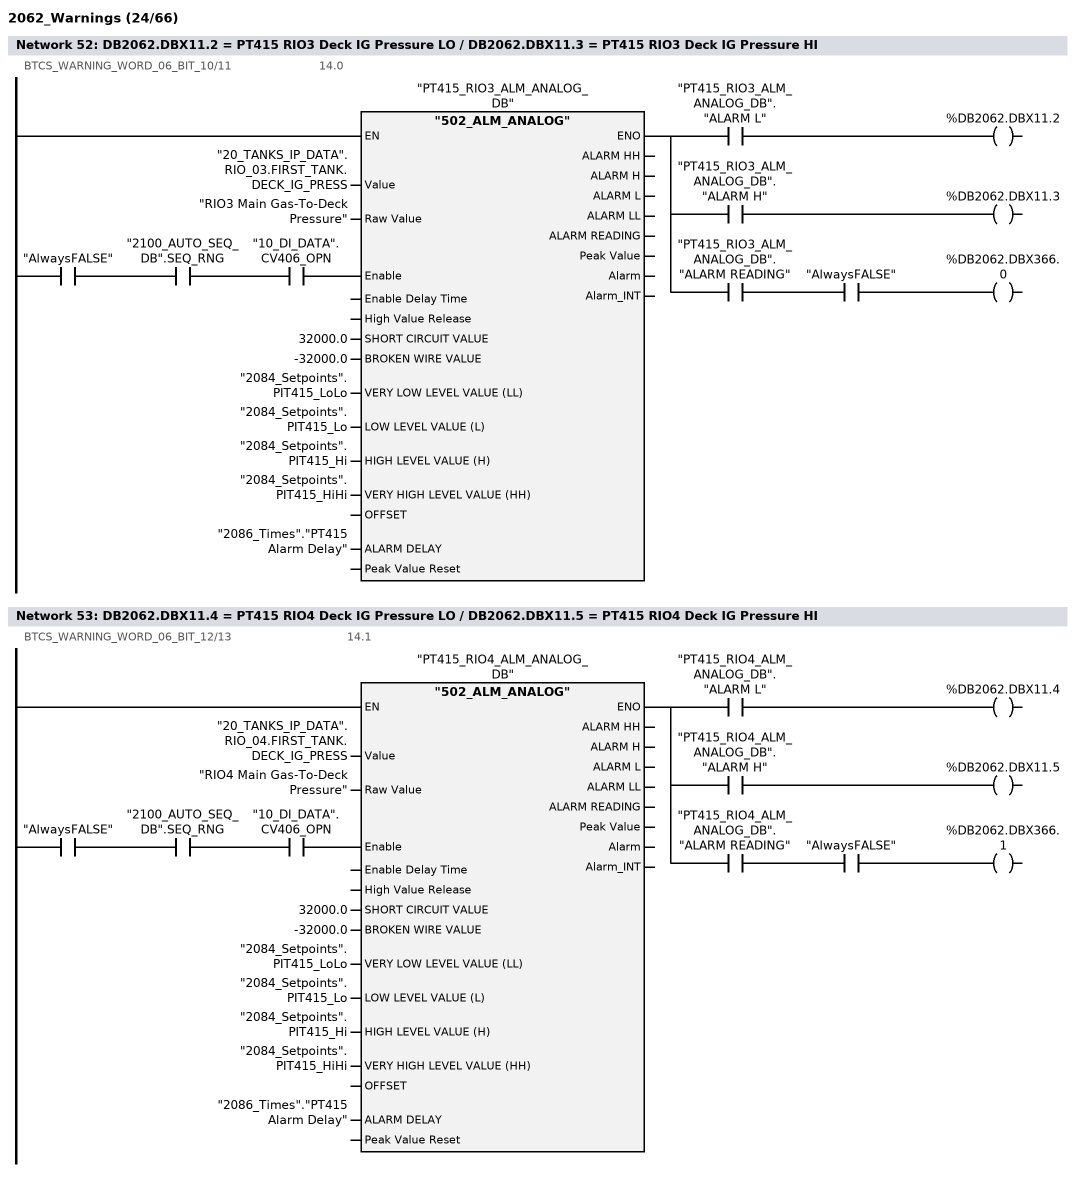
   RUNG wire#powerrail
      "PT415_RIO3_ALM_ANALOG_DB"(Enable := wire#w1, Value := "20_TANKS_IP_DATA".RIO_03.FIRST_TANK.DECK_IG_PRESS, "Raw Value" := "RIO3 Main Gas-To-Deck Pressure", "Enable Delay Time" :=, "High Value Release" :=, "SHORT CIRCUIT VALUE" := 32000.0, "BROKEN WIRE VALUE" := -32000.0, "VERY LOW LEVEL VALUE (LL)" := "2084_Setpoints".PIT415_LoLo, "LOW LEVEL VALUE (L)" := "2084_Setpoints".PIT415_Lo, "HIGH LEVEL VALUE (H)" := "2084_Setpoints".PIT415_Hi, "VERY HIGH LEVEL VALUE (HH)" := "2084_Setpoints".PIT415_HiHi, OFFSET :=, "ALARM DELAY" := "2086_Times"."PT415 Alarm Delay", "Peak Value Reset" :=, "ALARM HH" =>, "ALARM H" =>, "ALARM L" =>, "ALARM LL" =>, "ALARM READING" =>, "Peak Value" =>, Alarm =>, Alarm_INT =>)
      wire#w2
      Contact( "PT415_RIO3_ALM_ANALOG_DB"."ALARM L" )
      Coil( %DB2062.DBX11.2 )
   END_RUNG
   RUNG wire#powerrail
      Contact( "AlwaysFALSE" )
      Contact( "2100_AUTO_SEQ_DB".SEQ_RNG )
      Contact( "10_DI_DATA".CV406_OPN )
   END_RUNG wire#w1
   RUNG wire#w2
      Contact( "PT415_RIO3_ALM_ANALOG_DB"."ALARM H" )
      Coil( %DB2062.DBX11.3 )
   END_RUNG
   RUNG wire#w2
      Contact( "PT415_RIO3_ALM_ANALOG_DB"."ALARM READING" )
      Contact( "AlwaysFALSE" )
      Coil( %DB2062.DBX366.0 )
   END_RUNG
   // the same network as SCL:
   "PT415_RIO3_ALM_ANALOG_DB"(Value := "20_TANKS_IP_DATA".RIO_03.FIRST_TANK.DECK_IG_PRESS,   // "502_ALM_ANALOG"
                           "Raw Value" := "RIO3 Main Gas-To-Deck Pressure",
                           Enable := "AlwaysFALSE" AND "2100_AUTO_SEQ_DB".SEQ_RNG AND "10_DI_DATA".CV406_OPN,
                           "SHORT CIRCUIT VALUE" := 32000.0,
                           "BROKEN WIRE VALUE" := -32000.0,
                           "VERY LOW LEVEL VALUE (LL)" := "2084_Setpoints".PIT415_LoLo,
                           "LOW LEVEL VALUE (L)" := "2084_Setpoints".PIT415_Lo,
                           "HIGH LEVEL VALUE (H)" := "2084_Setpoints".PIT415_Hi,
                           "VERY HIGH LEVEL VALUE (HH)" := "2084_Setpoints".PIT415_HiHi,
                           "ALARM DELAY" := "2086_Times"."PT415 Alarm Delay",
                           ENO => #_w1);
   %DB2062.DBX11.2 := #_w1 AND "PT415_RIO3_ALM_ANALOG_DB"."ALARM L";
   %DB2062.DBX11.3 := #_w1 AND "PT415_RIO3_ALM_ANALOG_DB"."ALARM H";
   %DB2062.DBX366.0 := #_w1 AND "PT415_RIO3_ALM_ANALOG_DB"."ALARM READING" AND "AlwaysFALSE";
END_REGION

REGION Network 53: DB2062.DBX11.4 = PT415 RIO4 Deck IG Pressure LO / DB2062.DBX11.5 = PT415 RIO4 Deck IG Pressure HI
   // BTCS_WARNING_WORD_06_BIT_12/13                                 14.1
   RUNG wire#powerrail
      "PT415_RIO4_ALM_ANALOG_DB"(Enable := wire#w1, Value := "20_TANKS_IP_DATA".RIO_04.FIRST_TANK.DECK_IG_PRESS, "Raw Value" := "RIO4 Main Gas-To-Deck Pressure", "Enable Delay Time" :=, "High Value Release" :=, "SHORT CIRCUIT VALUE" := 32000.0, "BROKEN WIRE VALUE" := -32000.0, "VERY LOW LEVEL VALUE (LL)" := "2084_Setpoints".PIT415_LoLo, "LOW LEVEL VALUE (L)" := "2084_Setpoints".PIT415_Lo, "HIGH LEVEL VALUE (H)" := "2084_Setpoints".PIT415_Hi, "VERY HIGH LEVEL VALUE (HH)" := "2084_Setpoints".PIT415_HiHi, OFFSET :=, "ALARM DELAY" := "2086_Times"."PT415 Alarm Delay", "Peak Value Reset" :=, "ALARM HH" =>, "ALARM H" =>, "ALARM L" =>, "ALARM LL" =>, "ALARM READING" =>, "Peak Value" =>, Alarm =>, Alarm_INT =>)
      wire#w2
      Contact( "PT415_RIO4_ALM_ANALOG_DB"."ALARM L" )
      Coil( %DB2062.DBX11.4 )
   END_RUNG
   RUNG wire#powerrail
      Contact( "AlwaysFALSE" )
      Contact( "2100_AUTO_SEQ_DB".SEQ_RNG )
      Contact( "10_DI_DATA".CV406_OPN )
   END_RUNG wire#w1
   RUNG wire#w2
      Contact( "PT415_RIO4_ALM_ANALOG_DB"."ALARM H" )
      Coil( %DB2062.DBX11.5 )
   END_RUNG
   RUNG wire#w2
      Contact( "PT415_RIO4_ALM_ANALOG_DB"."ALARM READING" )
      Contact( "AlwaysFALSE" )
      Coil( %DB2062.DBX366.1 )
   END_RUNG
   // the same network as SCL:
   "PT415_RIO4_ALM_ANALOG_DB"(Value := "20_TANKS_IP_DATA".RIO_04.FIRST_TANK.DECK_IG_PRESS,   // "502_ALM_ANALOG"
                           "Raw Value" := "RIO4 Main Gas-To-Deck Pressure",
                           Enable := "AlwaysFALSE" AND "2100_AUTO_SEQ_DB".SEQ_RNG AND "10_DI_DATA".CV406_OPN,
                           "SHORT CIRCUIT VALUE" := 32000.0,
                           "BROKEN WIRE VALUE" := -32000.0,
                           "VERY LOW LEVEL VALUE (LL)" := "2084_Setpoints".PIT415_LoLo,
                           "LOW LEVEL VALUE (L)" := "2084_Setpoints".PIT415_Lo,
                           "HIGH LEVEL VALUE (H)" := "2084_Setpoints".PIT415_Hi,
                           "VERY HIGH LEVEL VALUE (HH)" := "2084_Setpoints".PIT415_HiHi,
                           "ALARM DELAY" := "2086_Times"."PT415 Alarm Delay",
                           ENO => #_w1);
   %DB2062.DBX11.4 := #_w1 AND "PT415_RIO4_ALM_ANALOG_DB"."ALARM L";
   %DB2062.DBX11.5 := #_w1 AND "PT415_RIO4_ALM_ANALOG_DB"."ALARM H";
   %DB2062.DBX366.1 := #_w1 AND "PT415_RIO4_ALM_ANALOG_DB"."ALARM READING" AND "AlwaysFALSE";
END_REGION

REGION Network 54: DB2062.DBX11.6 = PT415 RIO5 Deck IG Pressure LO / DB2062.DBX11.7 = PT415 RIO5 Deck IG Pressure HI
   // BTCS_WARNING_WORD_06_BIT_14/15                               14.2
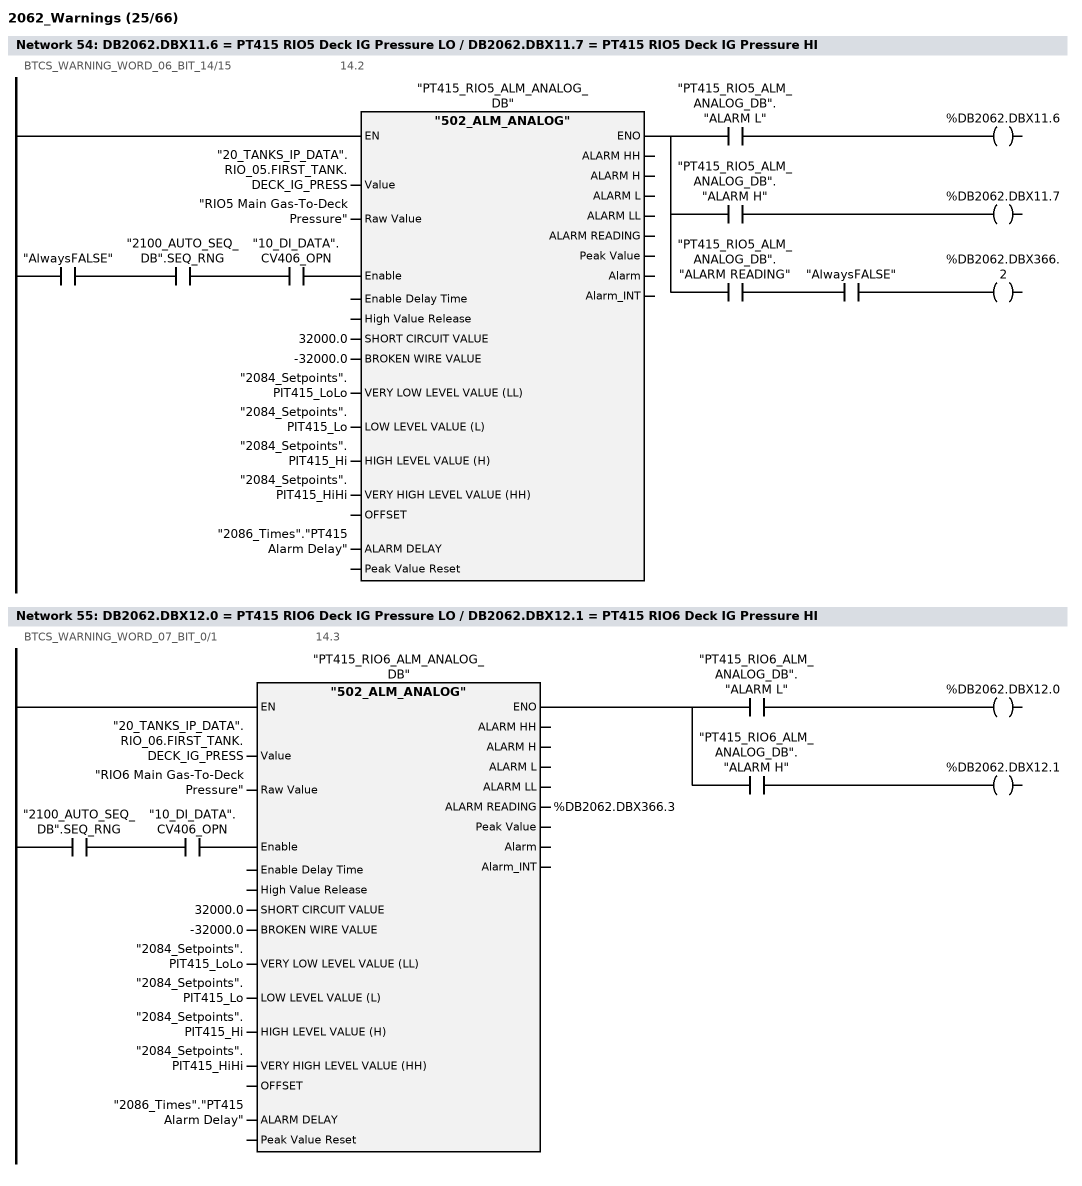
   RUNG wire#powerrail
      "PT415_RIO5_ALM_ANALOG_DB"(Enable := wire#w1, Value := "20_TANKS_IP_DATA".RIO_05.FIRST_TANK.DECK_IG_PRESS, "Raw Value" := "RIO5 Main Gas-To-Deck Pressure", "Enable Delay Time" :=, "High Value Release" :=, "SHORT CIRCUIT VALUE" := 32000.0, "BROKEN WIRE VALUE" := -32000.0, "VERY LOW LEVEL VALUE (LL)" := "2084_Setpoints".PIT415_LoLo, "LOW LEVEL VALUE (L)" := "2084_Setpoints".PIT415_Lo, "HIGH LEVEL VALUE (H)" := "2084_Setpoints".PIT415_Hi, "VERY HIGH LEVEL VALUE (HH)" := "2084_Setpoints".PIT415_HiHi, OFFSET :=, "ALARM DELAY" := "2086_Times"."PT415 Alarm Delay", "Peak Value Reset" :=, "ALARM HH" =>, "ALARM H" =>, "ALARM L" =>, "ALARM LL" =>, "ALARM READING" =>, "Peak Value" =>, Alarm =>, Alarm_INT =>)
      wire#w2
      Contact( "PT415_RIO5_ALM_ANALOG_DB"."ALARM L" )
      Coil( %DB2062.DBX11.6 )
   END_RUNG
   RUNG wire#powerrail
      Contact( "AlwaysFALSE" )
      Contact( "2100_AUTO_SEQ_DB".SEQ_RNG )
      Contact( "10_DI_DATA".CV406_OPN )
   END_RUNG wire#w1
   RUNG wire#w2
      Contact( "PT415_RIO5_ALM_ANALOG_DB"."ALARM H" )
      Coil( %DB2062.DBX11.7 )
   END_RUNG
   RUNG wire#w2
      Contact( "PT415_RIO5_ALM_ANALOG_DB"."ALARM READING" )
      Contact( "AlwaysFALSE" )
      Coil( %DB2062.DBX366.2 )
   END_RUNG
   // the same network as SCL:
   "PT415_RIO5_ALM_ANALOG_DB"(Value := "20_TANKS_IP_DATA".RIO_05.FIRST_TANK.DECK_IG_PRESS,   // "502_ALM_ANALOG"
                           "Raw Value" := "RIO5 Main Gas-To-Deck Pressure",
                           Enable := "AlwaysFALSE" AND "2100_AUTO_SEQ_DB".SEQ_RNG AND "10_DI_DATA".CV406_OPN,
                           "SHORT CIRCUIT VALUE" := 32000.0,
                           "BROKEN WIRE VALUE" := -32000.0,
                           "VERY LOW LEVEL VALUE (LL)" := "2084_Setpoints".PIT415_LoLo,
                           "LOW LEVEL VALUE (L)" := "2084_Setpoints".PIT415_Lo,
                           "HIGH LEVEL VALUE (H)" := "2084_Setpoints".PIT415_Hi,
                           "VERY HIGH LEVEL VALUE (HH)" := "2084_Setpoints".PIT415_HiHi,
                           "ALARM DELAY" := "2086_Times"."PT415 Alarm Delay",
                           ENO => #_w1);
   %DB2062.DBX11.6 := #_w1 AND "PT415_RIO5_ALM_ANALOG_DB"."ALARM L";
   %DB2062.DBX11.7 := #_w1 AND "PT415_RIO5_ALM_ANALOG_DB"."ALARM H";
   %DB2062.DBX366.2 := #_w1 AND "PT415_RIO5_ALM_ANALOG_DB"."ALARM READING" AND "AlwaysFALSE";
END_REGION

REGION Network 55: DB2062.DBX12.0 = PT415 RIO6 Deck IG Pressure LO / DB2062.DBX12.1 = PT415 RIO6 Deck IG Pressure HI
   // BTCS_WARNING_WORD_07_BIT_0/1                            14.3
   RUNG wire#powerrail
      "PT415_RIO6_ALM_ANALOG_DB"(Enable := wire#w1, Value := "20_TANKS_IP_DATA".RIO_06.FIRST_TANK.DECK_IG_PRESS, "Raw Value" := "RIO6 Main Gas-To-Deck Pressure", "Enable Delay Time" :=, "High Value Release" :=, "SHORT CIRCUIT VALUE" := 32000.0, "BROKEN WIRE VALUE" := -32000.0, "VERY LOW LEVEL VALUE (LL)" := "2084_Setpoints".PIT415_LoLo, "LOW LEVEL VALUE (L)" := "2084_Setpoints".PIT415_Lo, "HIGH LEVEL VALUE (H)" := "2084_Setpoints".PIT415_Hi, "VERY HIGH LEVEL VALUE (HH)" := "2084_Setpoints".PIT415_HiHi, OFFSET :=, "ALARM DELAY" := "2086_Times"."PT415 Alarm Delay", "Peak Value Reset" :=, "ALARM HH" =>, "ALARM H" =>, "ALARM L" =>, "ALARM LL" =>, "ALARM READING" => %DB2062.DBX366.3, "Peak Value" =>, Alarm =>, Alarm_INT =>)
      wire#w2
      Contact( "PT415_RIO6_ALM_ANALOG_DB"."ALARM L" )
      Coil( %DB2062.DBX12.0 )
   END_RUNG
   RUNG wire#powerrail
      Contact( "2100_AUTO_SEQ_DB".SEQ_RNG )
      Contact( "10_DI_DATA".CV406_OPN )
   END_RUNG wire#w1
   RUNG wire#w2
      Contact( "PT415_RIO6_ALM_ANALOG_DB"."ALARM H" )
      Coil( %DB2062.DBX12.1 )
   END_RUNG
   // the same network as SCL:
   "PT415_RIO6_ALM_ANALOG_DB"(Value := "20_TANKS_IP_DATA".RIO_06.FIRST_TANK.DECK_IG_PRESS,   // "502_ALM_ANALOG"
                           "Raw Value" := "RIO6 Main Gas-To-Deck Pressure",
                           Enable := "2100_AUTO_SEQ_DB".SEQ_RNG AND "10_DI_DATA".CV406_OPN,
                           "SHORT CIRCUIT VALUE" := 32000.0,
                           "BROKEN WIRE VALUE" := -32000.0,
                           "VERY LOW LEVEL VALUE (LL)" := "2084_Setpoints".PIT415_LoLo,
                           "LOW LEVEL VALUE (L)" := "2084_Setpoints".PIT415_Lo,
                           "HIGH LEVEL VALUE (H)" := "2084_Setpoints".PIT415_Hi,
                           "VERY HIGH LEVEL VALUE (HH)" := "2084_Setpoints".PIT415_HiHi,
                           "ALARM DELAY" := "2086_Times"."PT415 Alarm Delay",
                           "ALARM READING" => %DB2062.DBX366.3,
                           ENO => #_w1);
   %DB2062.DBX12.0 := #_w1 AND "PT415_RIO6_ALM_ANALOG_DB"."ALARM L";
   %DB2062.DBX12.1 := #_w1 AND "PT415_RIO6_ALM_ANALOG_DB"."ALARM H";
END_REGION

REGION Network 56: DB2062.DBX14.0 = PT415 RIO7 Deck IG Pressure LO / DB2062.DBX14.1 = PT415 RIO7 Deck IG Pressure HI
   // BTCS_WARNING_WORD_08_BIT_0/1                        14.4
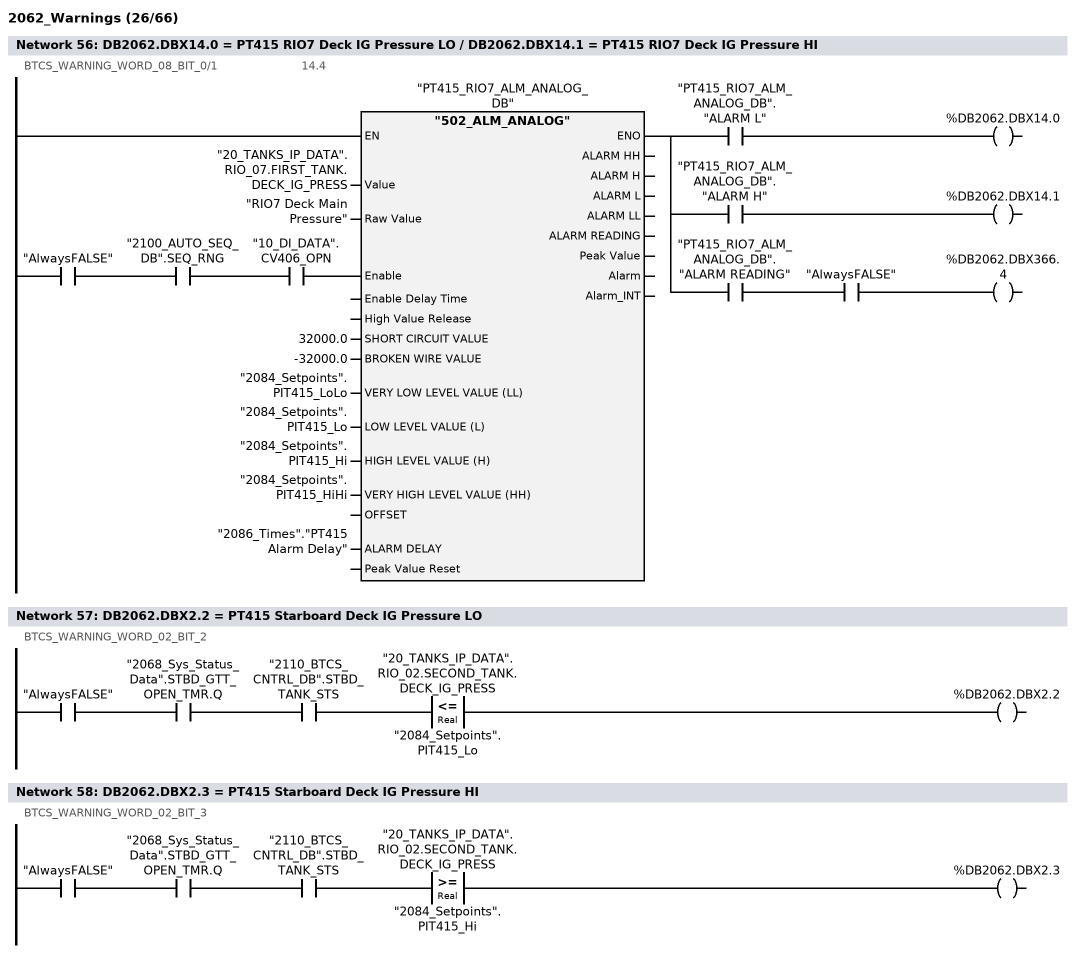
   RUNG wire#powerrail
      "PT415_RIO7_ALM_ANALOG_DB"(Enable := wire#w1, Value := "20_TANKS_IP_DATA".RIO_07.FIRST_TANK.DECK_IG_PRESS, "Raw Value" := "RIO7 Deck Main Pressure", "Enable Delay Time" :=, "High Value Release" :=, "SHORT CIRCUIT VALUE" := 32000.0, "BROKEN WIRE VALUE" := -32000.0, "VERY LOW LEVEL VALUE (LL)" := "2084_Setpoints".PIT415_LoLo, "LOW LEVEL VALUE (L)" := "2084_Setpoints".PIT415_Lo, "HIGH LEVEL VALUE (H)" := "2084_Setpoints".PIT415_Hi, "VERY HIGH LEVEL VALUE (HH)" := "2084_Setpoints".PIT415_HiHi, OFFSET :=, "ALARM DELAY" := "2086_Times"."PT415 Alarm Delay", "Peak Value Reset" :=, "ALARM HH" =>, "ALARM H" =>, "ALARM L" =>, "ALARM LL" =>, "ALARM READING" =>, "Peak Value" =>, Alarm =>, Alarm_INT =>)
      wire#w2
      Contact( "PT415_RIO7_ALM_ANALOG_DB"."ALARM L" )
      Coil( %DB2062.DBX14.0 )
   END_RUNG
   RUNG wire#powerrail
      Contact( "AlwaysFALSE" )
      Contact( "2100_AUTO_SEQ_DB".SEQ_RNG )
      Contact( "10_DI_DATA".CV406_OPN )
   END_RUNG wire#w1
   RUNG wire#w2
      Contact( "PT415_RIO7_ALM_ANALOG_DB"."ALARM H" )
      Coil( %DB2062.DBX14.1 )
   END_RUNG
   RUNG wire#w2
      Contact( "PT415_RIO7_ALM_ANALOG_DB"."ALARM READING" )
      Contact( "AlwaysFALSE" )
      Coil( %DB2062.DBX366.4 )
   END_RUNG
   // the same network as SCL:
   "PT415_RIO7_ALM_ANALOG_DB"(Value := "20_TANKS_IP_DATA".RIO_07.FIRST_TANK.DECK_IG_PRESS,   // "502_ALM_ANALOG"
                           "Raw Value" := "RIO7 Deck Main Pressure",
                           Enable := "AlwaysFALSE" AND "2100_AUTO_SEQ_DB".SEQ_RNG AND "10_DI_DATA".CV406_OPN,
                           "SHORT CIRCUIT VALUE" := 32000.0,
                           "BROKEN WIRE VALUE" := -32000.0,
                           "VERY LOW LEVEL VALUE (LL)" := "2084_Setpoints".PIT415_LoLo,
                           "LOW LEVEL VALUE (L)" := "2084_Setpoints".PIT415_Lo,
                           "HIGH LEVEL VALUE (H)" := "2084_Setpoints".PIT415_Hi,
                           "VERY HIGH LEVEL VALUE (HH)" := "2084_Setpoints".PIT415_HiHi,
                           "ALARM DELAY" := "2086_Times"."PT415 Alarm Delay",
                           ENO => #_w1);
   %DB2062.DBX14.0 := #_w1 AND "PT415_RIO7_ALM_ANALOG_DB"."ALARM L";
   %DB2062.DBX14.1 := #_w1 AND "PT415_RIO7_ALM_ANALOG_DB"."ALARM H";
   %DB2062.DBX366.4 := #_w1 AND "PT415_RIO7_ALM_ANALOG_DB"."ALARM READING" AND "AlwaysFALSE";
END_REGION

REGION Network 57: DB2062.DBX2.2 = PT415 Starboard Deck IG Pressure LO
   // BTCS_WARNING_WORD_02_BIT_2
   RUNG wire#powerrail
      Contact( "AlwaysFALSE" )
      Contact( "2068_Sys_Status_Data".STBD_GTT_OPEN_TMR.Q )
      Contact( "2110_BTCS_CNTRL_DB".STBD_TANK_STS )
      { S7_Templates := "SrcType := Real" } LE_Contact(in1 := "20_TANKS_IP_DATA".RIO_02.SECOND_TANK.DECK_IG_PRESS, in2 := "2084_Setpoints".PIT415_Lo)
      Coil( %DB2062.DBX2.2 )
   END_RUNG
   // the same network as SCL:
   %DB2062.DBX2.2 := "AlwaysFALSE" AND "2068_Sys_Status_Data".STBD_GTT_OPEN_TMR.Q AND "2110_BTCS_CNTRL_DB".STBD_TANK_STS AND ("20_TANKS_IP_DATA".RIO_02.SECOND_TANK.DECK_IG_PRESS <= "2084_Setpoints".PIT415_Lo);
END_REGION

REGION Network 58: DB2062.DBX2.3 = PT415 Starboard Deck IG Pressure HI
   // BTCS_WARNING_WORD_02_BIT_3
   RUNG wire#powerrail
      Contact( "AlwaysFALSE" )
      Contact( "2068_Sys_Status_Data".STBD_GTT_OPEN_TMR.Q )
      Contact( "2110_BTCS_CNTRL_DB".STBD_TANK_STS )
      { S7_Templates := "SrcType := Real" } GE_Contact(in1 := "20_TANKS_IP_DATA".RIO_02.SECOND_TANK.DECK_IG_PRESS, in2 := "2084_Setpoints".PIT415_Hi)
      Coil( %DB2062.DBX2.3 )
   END_RUNG
   // the same network as SCL:
   %DB2062.DBX2.3 := "AlwaysFALSE" AND "2068_Sys_Status_Data".STBD_GTT_OPEN_TMR.Q AND "2110_BTCS_CNTRL_DB".STBD_TANK_STS AND ("20_TANKS_IP_DATA".RIO_02.SECOND_TANK.DECK_IG_PRESS >= "2084_Setpoints".PIT415_Hi);
END_REGION

REGION Network 60: DB2062.DBX12.2/3 = PIT424 RIO1 Tank Pressure LO/HI
   // BTCS_WARNING_WORD_07_BIT_2/3                          14.5
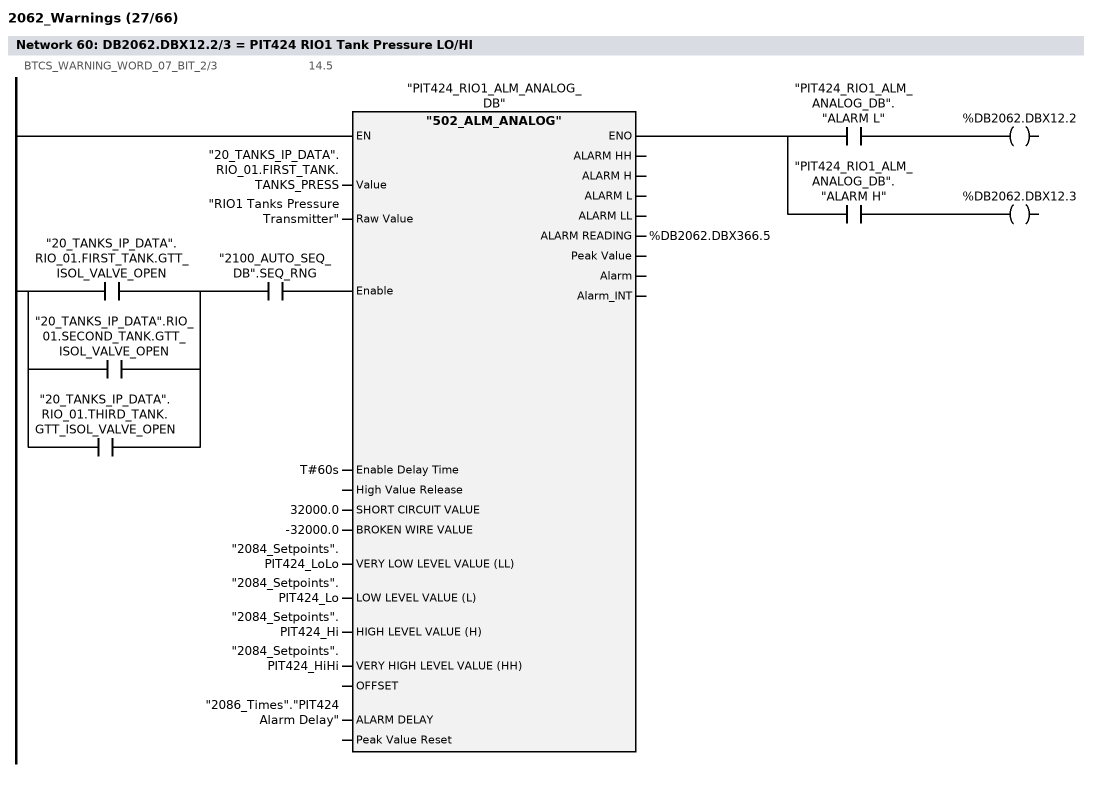
   RUNG wire#powerrail
      "PIT424_RIO1_ALM_ANALOG_DB"(Enable := wire#w2, Value := "20_TANKS_IP_DATA".RIO_01.FIRST_TANK.TANKS_PRESS, "Raw Value" := "RIO1 Tanks Pressure Transmitter", "Enable Delay Time" := T#60s, "High Value Release" :=, "SHORT CIRCUIT VALUE" := 32000.0, "BROKEN WIRE VALUE" := -32000.0, "VERY LOW LEVEL VALUE (LL)" := "2084_Setpoints".PIT424_LoLo, "LOW LEVEL VALUE (L)" := "2084_Setpoints".PIT424_Lo, "HIGH LEVEL VALUE (H)" := "2084_Setpoints".PIT424_Hi, "VERY HIGH LEVEL VALUE (HH)" := "2084_Setpoints".PIT424_HiHi, OFFSET :=, "ALARM DELAY" := "2086_Times"."PIT424 Alarm Delay", "Peak Value Reset" :=, "ALARM HH" =>, "ALARM H" =>, "ALARM L" =>, "ALARM LL" =>, "ALARM READING" => %DB2062.DBX366.5, "Peak Value" =>, Alarm =>, Alarm_INT =>)
      wire#w3
      Contact( "PIT424_RIO1_ALM_ANALOG_DB"."ALARM L" )
      Coil( %DB2062.DBX12.2 )
   END_RUNG
   RUNG wire#powerrail
      Contact( "20_TANKS_IP_DATA".RIO_01.FIRST_TANK.GTT_ISOL_VALVE_OPEN )
      wire#w1
      Contact( "2100_AUTO_SEQ_DB".SEQ_RNG )
   END_RUNG wire#w2
   RUNG wire#powerrail
      Contact( "20_TANKS_IP_DATA".RIO_01.SECOND_TANK.GTT_ISOL_VALVE_OPEN )
   END_RUNG wire#w1
   RUNG wire#powerrail
      Contact( "20_TANKS_IP_DATA".RIO_01.THIRD_TANK.GTT_ISOL_VALVE_OPEN )
   END_RUNG wire#w1
   RUNG wire#w3
      Contact( "PIT424_RIO1_ALM_ANALOG_DB"."ALARM H" )
      Coil( %DB2062.DBX12.3 )
   END_RUNG
   // the same network as SCL:
   "PIT424_RIO1_ALM_ANALOG_DB"(Value := "20_TANKS_IP_DATA".RIO_01.FIRST_TANK.TANKS_PRESS,   // "502_ALM_ANALOG"
                           "Raw Value" := "RIO1 Tanks Pressure Transmitter",
                           Enable := ("20_TANKS_IP_DATA".RIO_01.FIRST_TANK.GTT_ISOL_VALVE_OPEN OR "20_TANKS_IP_DATA".RIO_01.SECOND_TANK.GTT_ISOL_VALVE_OPEN OR "20_TANKS_IP_DATA".RIO_01.THIRD_TANK.GTT_ISOL_VALVE_OPEN) AND "2100_AUTO_SEQ_DB".SEQ_RNG,
                           "Enable Delay Time" := T#60s,
                           "SHORT CIRCUIT VALUE" := 32000.0,
                           "BROKEN WIRE VALUE" := -32000.0,
                           "VERY LOW LEVEL VALUE (LL)" := "2084_Setpoints".PIT424_LoLo,
                           "LOW LEVEL VALUE (L)" := "2084_Setpoints".PIT424_Lo,
                           "HIGH LEVEL VALUE (H)" := "2084_Setpoints".PIT424_Hi,
                           "VERY HIGH LEVEL VALUE (HH)" := "2084_Setpoints".PIT424_HiHi,
                           "ALARM DELAY" := "2086_Times"."PIT424 Alarm Delay",
                           "ALARM READING" => %DB2062.DBX366.5,
                           ENO => #_w1);
   %DB2062.DBX12.2 := #_w1 AND "PIT424_RIO1_ALM_ANALOG_DB"."ALARM L";
   %DB2062.DBX12.3 := #_w1 AND "PIT424_RIO1_ALM_ANALOG_DB"."ALARM H";
END_REGION

REGION Network 61: DB2062.DBX2.4/5 = PIT424 RIO2 Tank Pressure LO/HI
   // BTCS_WARNING_WORD_02_BIT_4                       14.6
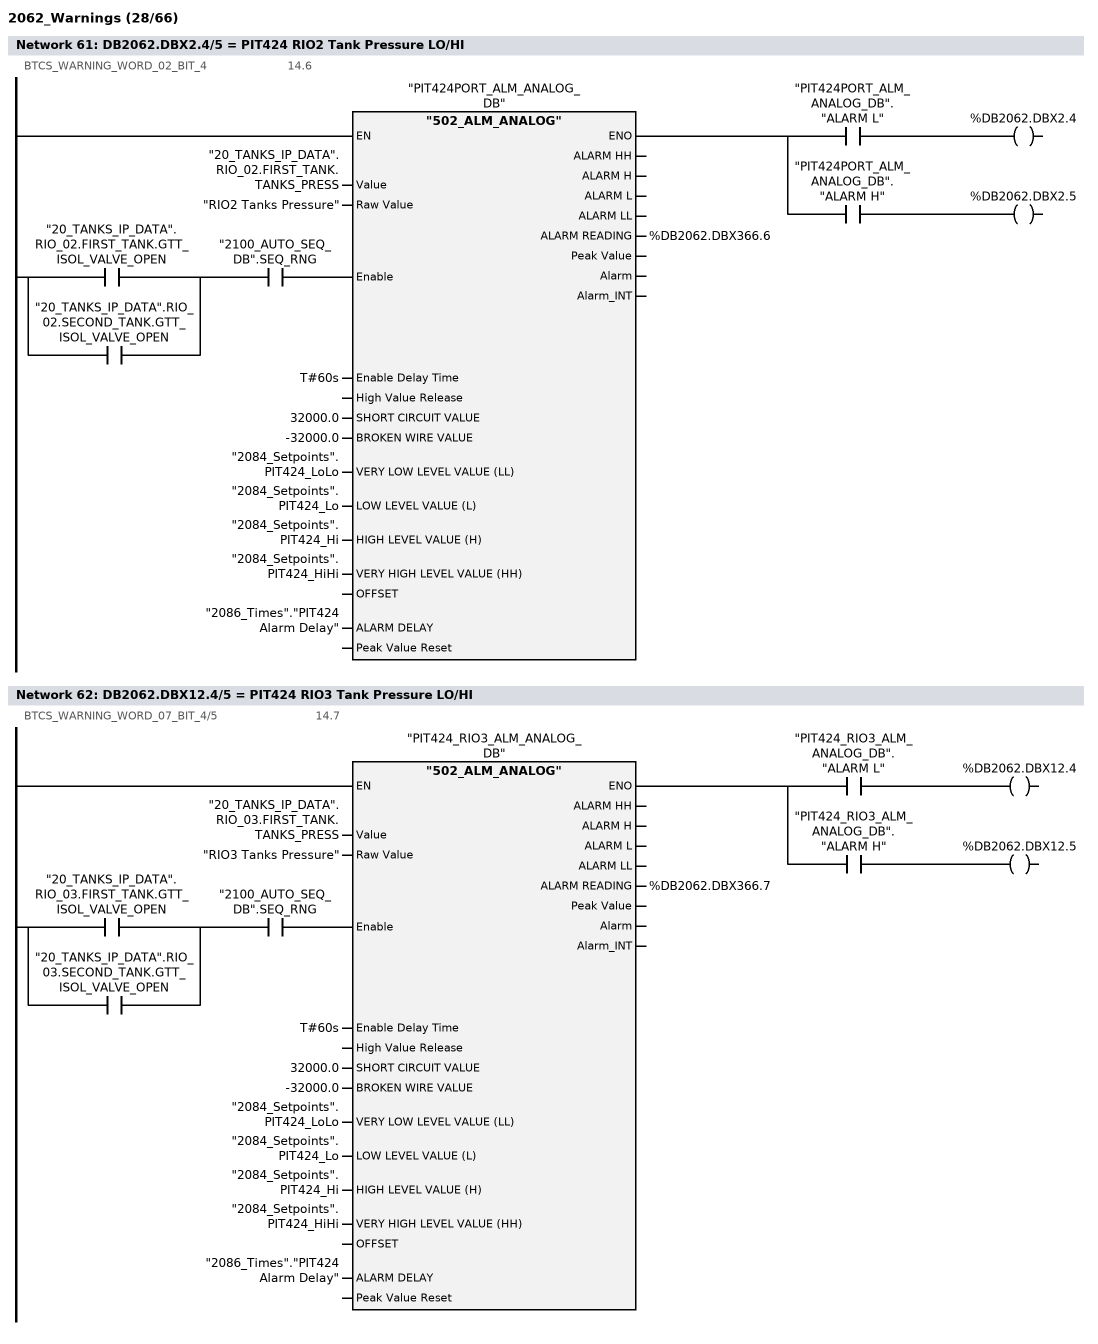
   RUNG wire#powerrail
      "PIT424PORT_ALM_ANALOG_DB"(Enable := wire#w2, Value := "20_TANKS_IP_DATA".RIO_02.FIRST_TANK.TANKS_PRESS, "Raw Value" := "RIO2 Tanks Pressure", "Enable Delay Time" := T#60s, "High Value Release" :=, "SHORT CIRCUIT VALUE" := 32000.0, "BROKEN WIRE VALUE" := -32000.0, "VERY LOW LEVEL VALUE (LL)" := "2084_Setpoints".PIT424_LoLo, "LOW LEVEL VALUE (L)" := "2084_Setpoints".PIT424_Lo, "HIGH LEVEL VALUE (H)" := "2084_Setpoints".PIT424_Hi, "VERY HIGH LEVEL VALUE (HH)" := "2084_Setpoints".PIT424_HiHi, OFFSET :=, "ALARM DELAY" := "2086_Times"."PIT424 Alarm Delay", "Peak Value Reset" :=, "ALARM HH" =>, "ALARM H" =>, "ALARM L" =>, "ALARM LL" =>, "ALARM READING" => %DB2062.DBX366.6, "Peak Value" =>, Alarm =>, Alarm_INT =>)
      wire#w3
      Contact( "PIT424PORT_ALM_ANALOG_DB"."ALARM L" )
      Coil( %DB2062.DBX2.4 )
   END_RUNG
   RUNG wire#powerrail
      Contact( "20_TANKS_IP_DATA".RIO_02.FIRST_TANK.GTT_ISOL_VALVE_OPEN )
      wire#w1
      Contact( "2100_AUTO_SEQ_DB".SEQ_RNG )
   END_RUNG wire#w2
   RUNG wire#powerrail
      Contact( "20_TANKS_IP_DATA".RIO_02.SECOND_TANK.GTT_ISOL_VALVE_OPEN )
   END_RUNG wire#w1
   RUNG wire#w3
      Contact( "PIT424PORT_ALM_ANALOG_DB"."ALARM H" )
      Coil( %DB2062.DBX2.5 )
   END_RUNG
   // the same network as SCL:
   "PIT424PORT_ALM_ANALOG_DB"(Value := "20_TANKS_IP_DATA".RIO_02.FIRST_TANK.TANKS_PRESS,   // "502_ALM_ANALOG"
                           "Raw Value" := "RIO2 Tanks Pressure",
                           Enable := ("20_TANKS_IP_DATA".RIO_02.FIRST_TANK.GTT_ISOL_VALVE_OPEN OR "20_TANKS_IP_DATA".RIO_02.SECOND_TANK.GTT_ISOL_VALVE_OPEN) AND "2100_AUTO_SEQ_DB".SEQ_RNG,
                           "Enable Delay Time" := T#60s,
                           "SHORT CIRCUIT VALUE" := 32000.0,
                           "BROKEN WIRE VALUE" := -32000.0,
                           "VERY LOW LEVEL VALUE (LL)" := "2084_Setpoints".PIT424_LoLo,
                           "LOW LEVEL VALUE (L)" := "2084_Setpoints".PIT424_Lo,
                           "HIGH LEVEL VALUE (H)" := "2084_Setpoints".PIT424_Hi,
                           "VERY HIGH LEVEL VALUE (HH)" := "2084_Setpoints".PIT424_HiHi,
                           "ALARM DELAY" := "2086_Times"."PIT424 Alarm Delay",
                           "ALARM READING" => %DB2062.DBX366.6,
                           ENO => #_w1);
   %DB2062.DBX2.4 := #_w1 AND "PIT424PORT_ALM_ANALOG_DB"."ALARM L";
   %DB2062.DBX2.5 := #_w1 AND "PIT424PORT_ALM_ANALOG_DB"."ALARM H";
END_REGION

REGION Network 62: DB2062.DBX12.4/5 = PIT424 RIO3 Tank Pressure LO/HI
   // BTCS_WARNING_WORD_07_BIT_4/5                            14.7
   RUNG wire#powerrail
      "PIT424_RIO3_ALM_ANALOG_DB"(Enable := wire#w2, Value := "20_TANKS_IP_DATA".RIO_03.FIRST_TANK.TANKS_PRESS, "Raw Value" := "RIO3 Tanks Pressure", "Enable Delay Time" := T#60s, "High Value Release" :=, "SHORT CIRCUIT VALUE" := 32000.0, "BROKEN WIRE VALUE" := -32000.0, "VERY LOW LEVEL VALUE (LL)" := "2084_Setpoints".PIT424_LoLo, "LOW LEVEL VALUE (L)" := "2084_Setpoints".PIT424_Lo, "HIGH LEVEL VALUE (H)" := "2084_Setpoints".PIT424_Hi, "VERY HIGH LEVEL VALUE (HH)" := "2084_Setpoints".PIT424_HiHi, OFFSET :=, "ALARM DELAY" := "2086_Times"."PIT424 Alarm Delay", "Peak Value Reset" :=, "ALARM HH" =>, "ALARM H" =>, "ALARM L" =>, "ALARM LL" =>, "ALARM READING" => %DB2062.DBX366.7, "Peak Value" =>, Alarm =>, Alarm_INT =>)
      wire#w3
      Contact( "PIT424_RIO3_ALM_ANALOG_DB"."ALARM L" )
      Coil( %DB2062.DBX12.4 )
   END_RUNG
   RUNG wire#powerrail
      Contact( "20_TANKS_IP_DATA".RIO_03.FIRST_TANK.GTT_ISOL_VALVE_OPEN )
      wire#w1
      Contact( "2100_AUTO_SEQ_DB".SEQ_RNG )
   END_RUNG wire#w2
   RUNG wire#powerrail
      Contact( "20_TANKS_IP_DATA".RIO_03.SECOND_TANK.GTT_ISOL_VALVE_OPEN )
   END_RUNG wire#w1
   RUNG wire#w3
      Contact( "PIT424_RIO3_ALM_ANALOG_DB"."ALARM H" )
      Coil( %DB2062.DBX12.5 )
   END_RUNG
   // the same network as SCL:
   "PIT424_RIO3_ALM_ANALOG_DB"(Value := "20_TANKS_IP_DATA".RIO_03.FIRST_TANK.TANKS_PRESS,   // "502_ALM_ANALOG"
                           "Raw Value" := "RIO3 Tanks Pressure",
                           Enable := ("20_TANKS_IP_DATA".RIO_03.FIRST_TANK.GTT_ISOL_VALVE_OPEN OR "20_TANKS_IP_DATA".RIO_03.SECOND_TANK.GTT_ISOL_VALVE_OPEN) AND "2100_AUTO_SEQ_DB".SEQ_RNG,
                           "Enable Delay Time" := T#60s,
                           "SHORT CIRCUIT VALUE" := 32000.0,
                           "BROKEN WIRE VALUE" := -32000.0,
                           "VERY LOW LEVEL VALUE (LL)" := "2084_Setpoints".PIT424_LoLo,
                           "LOW LEVEL VALUE (L)" := "2084_Setpoints".PIT424_Lo,
                           "HIGH LEVEL VALUE (H)" := "2084_Setpoints".PIT424_Hi,
                           "VERY HIGH LEVEL VALUE (HH)" := "2084_Setpoints".PIT424_HiHi,
                           "ALARM DELAY" := "2086_Times"."PIT424 Alarm Delay",
                           "ALARM READING" => %DB2062.DBX366.7,
                           ENO => #_w1);
   %DB2062.DBX12.4 := #_w1 AND "PIT424_RIO3_ALM_ANALOG_DB"."ALARM L";
   %DB2062.DBX12.5 := #_w1 AND "PIT424_RIO3_ALM_ANALOG_DB"."ALARM H";
END_REGION

REGION Network 63: DB2062.DBX12.6/7 = PIT424 RIO4 Tank Pressure LO/HI
   // BTCS_WARNING_WORD_07_BIT_6/7                           14.8
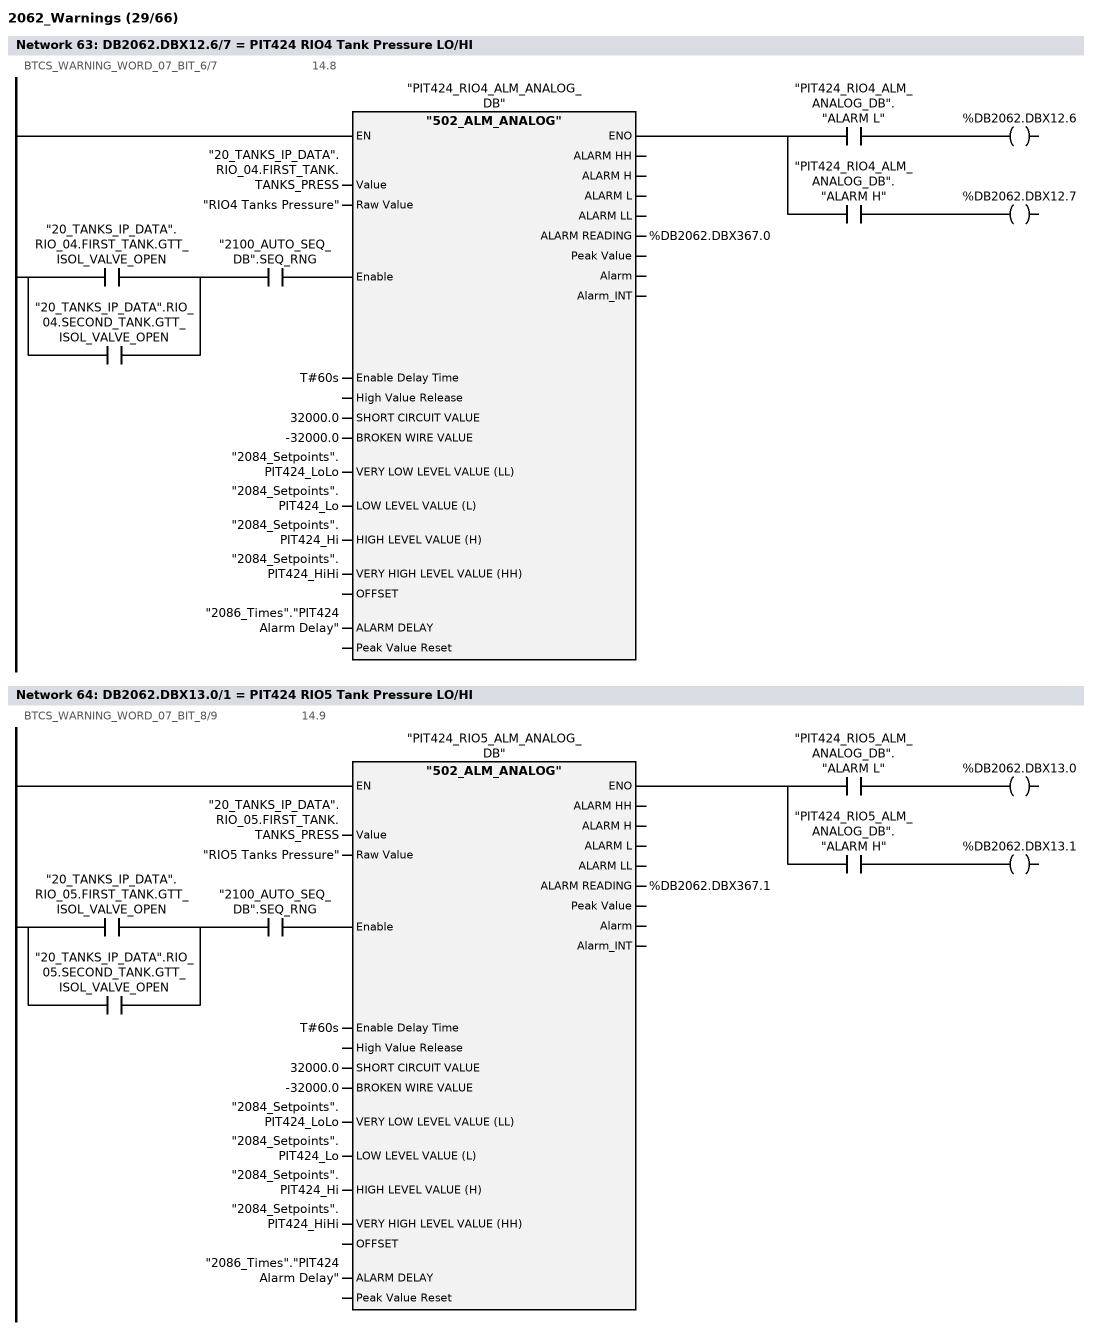
   RUNG wire#powerrail
      "PIT424_RIO4_ALM_ANALOG_DB"(Enable := wire#w2, Value := "20_TANKS_IP_DATA".RIO_04.FIRST_TANK.TANKS_PRESS, "Raw Value" := "RIO4 Tanks Pressure", "Enable Delay Time" := T#60s, "High Value Release" :=, "SHORT CIRCUIT VALUE" := 32000.0, "BROKEN WIRE VALUE" := -32000.0, "VERY LOW LEVEL VALUE (LL)" := "2084_Setpoints".PIT424_LoLo, "LOW LEVEL VALUE (L)" := "2084_Setpoints".PIT424_Lo, "HIGH LEVEL VALUE (H)" := "2084_Setpoints".PIT424_Hi, "VERY HIGH LEVEL VALUE (HH)" := "2084_Setpoints".PIT424_HiHi, OFFSET :=, "ALARM DELAY" := "2086_Times"."PIT424 Alarm Delay", "Peak Value Reset" :=, "ALARM HH" =>, "ALARM H" =>, "ALARM L" =>, "ALARM LL" =>, "ALARM READING" => %DB2062.DBX367.0, "Peak Value" =>, Alarm =>, Alarm_INT =>)
      wire#w3
      Contact( "PIT424_RIO4_ALM_ANALOG_DB"."ALARM L" )
      Coil( %DB2062.DBX12.6 )
   END_RUNG
   RUNG wire#powerrail
      Contact( "20_TANKS_IP_DATA".RIO_04.FIRST_TANK.GTT_ISOL_VALVE_OPEN )
      wire#w1
      Contact( "2100_AUTO_SEQ_DB".SEQ_RNG )
   END_RUNG wire#w2
   RUNG wire#powerrail
      Contact( "20_TANKS_IP_DATA".RIO_04.SECOND_TANK.GTT_ISOL_VALVE_OPEN )
   END_RUNG wire#w1
   RUNG wire#w3
      Contact( "PIT424_RIO4_ALM_ANALOG_DB"."ALARM H" )
      Coil( %DB2062.DBX12.7 )
   END_RUNG
   // the same network as SCL:
   "PIT424_RIO4_ALM_ANALOG_DB"(Value := "20_TANKS_IP_DATA".RIO_04.FIRST_TANK.TANKS_PRESS,   // "502_ALM_ANALOG"
                           "Raw Value" := "RIO4 Tanks Pressure",
                           Enable := ("20_TANKS_IP_DATA".RIO_04.FIRST_TANK.GTT_ISOL_VALVE_OPEN OR "20_TANKS_IP_DATA".RIO_04.SECOND_TANK.GTT_ISOL_VALVE_OPEN) AND "2100_AUTO_SEQ_DB".SEQ_RNG,
                           "Enable Delay Time" := T#60s,
                           "SHORT CIRCUIT VALUE" := 32000.0,
                           "BROKEN WIRE VALUE" := -32000.0,
                           "VERY LOW LEVEL VALUE (LL)" := "2084_Setpoints".PIT424_LoLo,
                           "LOW LEVEL VALUE (L)" := "2084_Setpoints".PIT424_Lo,
                           "HIGH LEVEL VALUE (H)" := "2084_Setpoints".PIT424_Hi,
                           "VERY HIGH LEVEL VALUE (HH)" := "2084_Setpoints".PIT424_HiHi,
                           "ALARM DELAY" := "2086_Times"."PIT424 Alarm Delay",
                           "ALARM READING" => %DB2062.DBX367.0,
                           ENO => #_w1);
   %DB2062.DBX12.6 := #_w1 AND "PIT424_RIO4_ALM_ANALOG_DB"."ALARM L";
   %DB2062.DBX12.7 := #_w1 AND "PIT424_RIO4_ALM_ANALOG_DB"."ALARM H";
END_REGION

REGION Network 64: DB2062.DBX13.0/1 = PIT424 RIO5 Tank Pressure LO/HI
   // BTCS_WARNING_WORD_07_BIT_8/9                        14.9
   RUNG wire#powerrail
      "PIT424_RIO5_ALM_ANALOG_DB"(Enable := wire#w2, Value := "20_TANKS_IP_DATA".RIO_05.FIRST_TANK.TANKS_PRESS, "Raw Value" := "RIO5 Tanks Pressure", "Enable Delay Time" := T#60s, "High Value Release" :=, "SHORT CIRCUIT VALUE" := 32000.0, "BROKEN WIRE VALUE" := -32000.0, "VERY LOW LEVEL VALUE (LL)" := "2084_Setpoints".PIT424_LoLo, "LOW LEVEL VALUE (L)" := "2084_Setpoints".PIT424_Lo, "HIGH LEVEL VALUE (H)" := "2084_Setpoints".PIT424_Hi, "VERY HIGH LEVEL VALUE (HH)" := "2084_Setpoints".PIT424_HiHi, OFFSET :=, "ALARM DELAY" := "2086_Times"."PIT424 Alarm Delay", "Peak Value Reset" :=, "ALARM HH" =>, "ALARM H" =>, "ALARM L" =>, "ALARM LL" =>, "ALARM READING" => %DB2062.DBX367.1, "Peak Value" =>, Alarm =>, Alarm_INT =>)
      wire#w3
      Contact( "PIT424_RIO5_ALM_ANALOG_DB"."ALARM L" )
      Coil( %DB2062.DBX13.0 )
   END_RUNG
   RUNG wire#powerrail
      Contact( "20_TANKS_IP_DATA".RIO_05.FIRST_TANK.GTT_ISOL_VALVE_OPEN )
      wire#w1
      Contact( "2100_AUTO_SEQ_DB".SEQ_RNG )
   END_RUNG wire#w2
   RUNG wire#powerrail
      Contact( "20_TANKS_IP_DATA".RIO_05.SECOND_TANK.GTT_ISOL_VALVE_OPEN )
   END_RUNG wire#w1
   RUNG wire#w3
      Contact( "PIT424_RIO5_ALM_ANALOG_DB"."ALARM H" )
      Coil( %DB2062.DBX13.1 )
   END_RUNG
   // the same network as SCL:
   "PIT424_RIO5_ALM_ANALOG_DB"(Value := "20_TANKS_IP_DATA".RIO_05.FIRST_TANK.TANKS_PRESS,   // "502_ALM_ANALOG"
                           "Raw Value" := "RIO5 Tanks Pressure",
                           Enable := ("20_TANKS_IP_DATA".RIO_05.FIRST_TANK.GTT_ISOL_VALVE_OPEN OR "20_TANKS_IP_DATA".RIO_05.SECOND_TANK.GTT_ISOL_VALVE_OPEN) AND "2100_AUTO_SEQ_DB".SEQ_RNG,
                           "Enable Delay Time" := T#60s,
                           "SHORT CIRCUIT VALUE" := 32000.0,
                           "BROKEN WIRE VALUE" := -32000.0,
                           "VERY LOW LEVEL VALUE (LL)" := "2084_Setpoints".PIT424_LoLo,
                           "LOW LEVEL VALUE (L)" := "2084_Setpoints".PIT424_Lo,
                           "HIGH LEVEL VALUE (H)" := "2084_Setpoints".PIT424_Hi,
                           "VERY HIGH LEVEL VALUE (HH)" := "2084_Setpoints".PIT424_HiHi,
                           "ALARM DELAY" := "2086_Times"."PIT424 Alarm Delay",
                           "ALARM READING" => %DB2062.DBX367.1,
                           ENO => #_w1);
   %DB2062.DBX13.0 := #_w1 AND "PIT424_RIO5_ALM_ANALOG_DB"."ALARM L";
   %DB2062.DBX13.1 := #_w1 AND "PIT424_RIO5_ALM_ANALOG_DB"."ALARM H";
END_REGION

REGION Network 65: DB2062.DBX13.2/3 = PIT424 RIO6 Tank Pressure LO/HI
   // BTCS_WARNING_WORD_07_BIT_10/11                             14.10